REGION Network 241: SAFE OUTPUT CARD FAULT
   RUNG wire#powerrail
      Contact( "reset" )
      { S7_Templates := "SrcType := Word" } EQ_Contact(in1 := "DB101_DB_SDC_FAULTS".Carrier_Fault[7], in2 := 122)
      Coil( "DB302_HMI_Faults".Carrier7_Faults_0.%X9 )
   END_RUNG
   // the same network as SCL:
   "DB302_HMI_Faults".Carrier7_Faults_0.%X9 := "reset" AND ("DB101_DB_SDC_FAULTS".Carrier_Fault[7] = 122);
END_REGION

REGION Network 242: STANDARD INPUT CARD FAULT
   RUNG wire#powerrail
      Contact( "reset" )
      { S7_Templates := "SrcType := Word" } EQ_Contact(in1 := "DB101_DB_SDC_FAULTS".Carrier_Fault[7], in2 := 123)
      Coil( "DB302_HMI_Faults".Carrier7_Faults_0.%X10 )
   END_RUNG
   // the same network as SCL:
   "DB302_HMI_Faults".Carrier7_Faults_0.%X10 := "reset" AND ("DB101_DB_SDC_FAULTS".Carrier_Fault[7] = 123);
END_REGION

REGION Network 243: STANDARD OUTPUT CARD FAULT
   RUNG wire#powerrail
      Contact( "reset" )
      { S7_Templates := "SrcType := Word" } EQ_Contact(in1 := "DB101_DB_SDC_FAULTS".Carrier_Fault[7], in2 := 124)
      Coil( "DB302_HMI_Faults".Carrier7_Faults_0.%X11 )
   END_RUNG
   // the same network as SCL:
   "DB302_HMI_Faults".Carrier7_Faults_0.%X11 := "reset" AND ("DB101_DB_SDC_FAULTS".Carrier_Fault[7] = 124);
END_REGION

REGION Network 244: CARRIER ENCODER POSITION FAULT
   RUNG wire#powerrail
      Contact( "reset" )
      { S7_Templates := "SrcType := Word" } EQ_Contact(in1 := "DB101_DB_SDC_FAULTS".Carrier_Fault[7], in2 := 131)
      Coil( "DB302_HMI_Faults".Carrier7_Faults_0.%X12 )
   END_RUNG
   // the same network as SCL:
   "DB302_HMI_Faults".Carrier7_Faults_0.%X12 := "reset" AND ("DB101_DB_SDC_FAULTS".Carrier_Fault[7] = 131);
END_REGION

REGION Network 245: CARRIER ENCODER INTERNAL ERROR
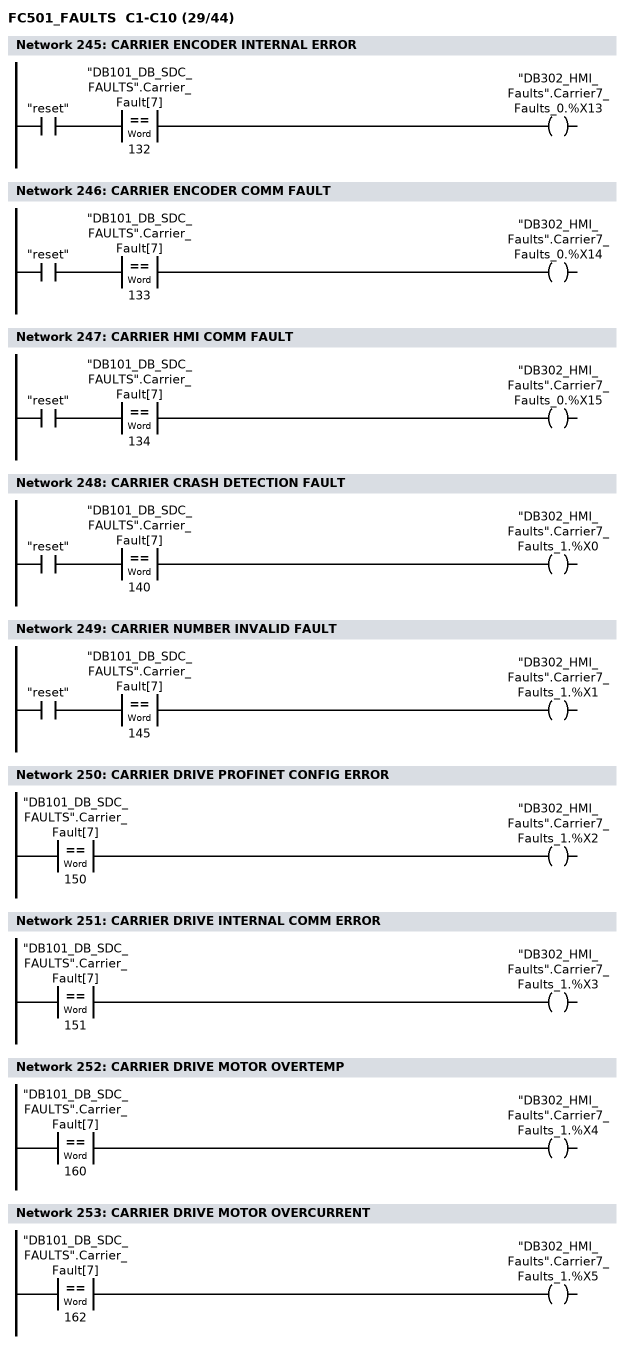
   RUNG wire#powerrail
      Contact( "reset" )
      { S7_Templates := "SrcType := Word" } EQ_Contact(in1 := "DB101_DB_SDC_FAULTS".Carrier_Fault[7], in2 := 132)
      Coil( "DB302_HMI_Faults".Carrier7_Faults_0.%X13 )
   END_RUNG
   // the same network as SCL:
   "DB302_HMI_Faults".Carrier7_Faults_0.%X13 := "reset" AND ("DB101_DB_SDC_FAULTS".Carrier_Fault[7] = 132);
END_REGION

REGION Network 246: CARRIER ENCODER COMM FAULT
   RUNG wire#powerrail
      Contact( "reset" )
      { S7_Templates := "SrcType := Word" } EQ_Contact(in1 := "DB101_DB_SDC_FAULTS".Carrier_Fault[7], in2 := 133)
      Coil( "DB302_HMI_Faults".Carrier7_Faults_0.%X14 )
   END_RUNG
   // the same network as SCL:
   "DB302_HMI_Faults".Carrier7_Faults_0.%X14 := "reset" AND ("DB101_DB_SDC_FAULTS".Carrier_Fault[7] = 133);
END_REGION

REGION Network 247: CARRIER HMI COMM FAULT
   RUNG wire#powerrail
      Contact( "reset" )
      { S7_Templates := "SrcType := Word" } EQ_Contact(in1 := "DB101_DB_SDC_FAULTS".Carrier_Fault[7], in2 := 134)
      Coil( "DB302_HMI_Faults".Carrier7_Faults_0.%X15 )
   END_RUNG
   // the same network as SCL:
   "DB302_HMI_Faults".Carrier7_Faults_0.%X15 := "reset" AND ("DB101_DB_SDC_FAULTS".Carrier_Fault[7] = 134);
END_REGION

REGION Network 248: CARRIER CRASH DETECTION FAULT
   RUNG wire#powerrail
      Contact( "reset" )
      { S7_Templates := "SrcType := Word" } EQ_Contact(in1 := "DB101_DB_SDC_FAULTS".Carrier_Fault[7], in2 := 140)
      Coil( "DB302_HMI_Faults".Carrier7_Faults_1.%X0 )
   END_RUNG
   // the same network as SCL:
   "DB302_HMI_Faults".Carrier7_Faults_1.%X0 := "reset" AND ("DB101_DB_SDC_FAULTS".Carrier_Fault[7] = 140);
END_REGION

REGION Network 249: CARRIER NUMBER INVALID FAULT
   RUNG wire#powerrail
      Contact( "reset" )
      { S7_Templates := "SrcType := Word" } EQ_Contact(in1 := "DB101_DB_SDC_FAULTS".Carrier_Fault[7], in2 := 145)
      Coil( "DB302_HMI_Faults".Carrier7_Faults_1.%X1 )
   END_RUNG
   // the same network as SCL:
   "DB302_HMI_Faults".Carrier7_Faults_1.%X1 := "reset" AND ("DB101_DB_SDC_FAULTS".Carrier_Fault[7] = 145);
END_REGION

REGION Network 250: CARRIER DRIVE PROFINET CONFIG ERROR
   RUNG wire#powerrail
      { S7_Templates := "SrcType := Word" } EQ_Contact(in1 := "DB101_DB_SDC_FAULTS".Carrier_Fault[7], in2 := 150)
      Coil( "DB302_HMI_Faults".Carrier7_Faults_1.%X2 )
   END_RUNG
   // the same network as SCL:
   "DB302_HMI_Faults".Carrier7_Faults_1.%X2 := "DB101_DB_SDC_FAULTS".Carrier_Fault[7] = 150;
END_REGION

REGION Network 251: CARRIER DRIVE INTERNAL COMM ERROR
   RUNG wire#powerrail
      { S7_Templates := "SrcType := Word" } EQ_Contact(in1 := "DB101_DB_SDC_FAULTS".Carrier_Fault[7], in2 := 151)
      Coil( "DB302_HMI_Faults".Carrier7_Faults_1.%X3 )
   END_RUNG
   // the same network as SCL:
   "DB302_HMI_Faults".Carrier7_Faults_1.%X3 := "DB101_DB_SDC_FAULTS".Carrier_Fault[7] = 151;
END_REGION

REGION Network 252: CARRIER DRIVE MOTOR OVERTEMP
   RUNG wire#powerrail
      { S7_Templates := "SrcType := Word" } EQ_Contact(in1 := "DB101_DB_SDC_FAULTS".Carrier_Fault[7], in2 := 160)
      Coil( "DB302_HMI_Faults".Carrier7_Faults_1.%X4 )
   END_RUNG
   // the same network as SCL:
   "DB302_HMI_Faults".Carrier7_Faults_1.%X4 := "DB101_DB_SDC_FAULTS".Carrier_Fault[7] = 160;
END_REGION

REGION Network 253: CARRIER DRIVE MOTOR OVERCURRENT
   RUNG wire#powerrail
      { S7_Templates := "SrcType := Word" } EQ_Contact(in1 := "DB101_DB_SDC_FAULTS".Carrier_Fault[7], in2 := 162)
      Coil( "DB302_HMI_Faults".Carrier7_Faults_1.%X5 )
   END_RUNG
   // the same network as SCL:
   "DB302_HMI_Faults".Carrier7_Faults_1.%X5 := "DB101_DB_SDC_FAULTS".Carrier_Fault[7] = 162;
END_REGION

REGION Network 254: CARRIER DRIVE INFEED OR POWER UNIT NOT READY
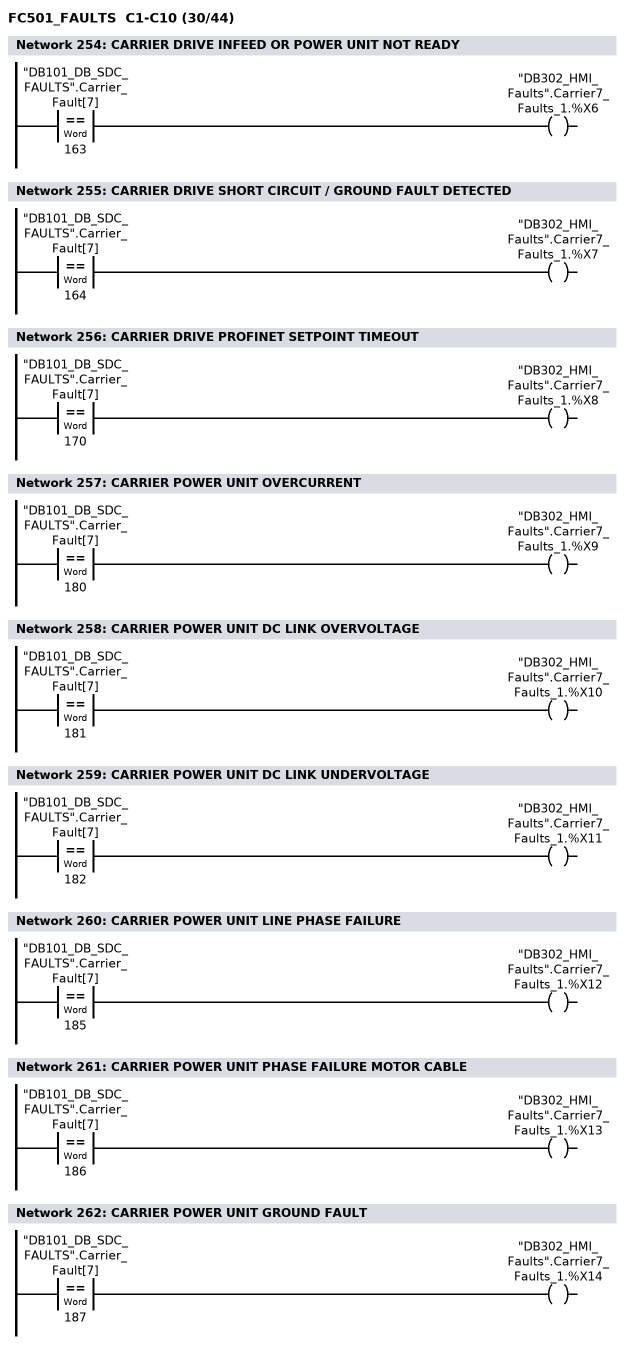
   RUNG wire#powerrail
      { S7_Templates := "SrcType := Word" } EQ_Contact(in1 := "DB101_DB_SDC_FAULTS".Carrier_Fault[7], in2 := 163)
      Coil( "DB302_HMI_Faults".Carrier7_Faults_1.%X6 )
   END_RUNG
   // the same network as SCL:
   "DB302_HMI_Faults".Carrier7_Faults_1.%X6 := "DB101_DB_SDC_FAULTS".Carrier_Fault[7] = 163;
END_REGION

REGION Network 255: CARRIER DRIVE SHORT CIRCUIT / GROUND FAULT DETECTED
   RUNG wire#powerrail
      { S7_Templates := "SrcType := Word" } EQ_Contact(in1 := "DB101_DB_SDC_FAULTS".Carrier_Fault[7], in2 := 164)
      Coil( "DB302_HMI_Faults".Carrier7_Faults_1.%X7 )
   END_RUNG
   // the same network as SCL:
   "DB302_HMI_Faults".Carrier7_Faults_1.%X7 := "DB101_DB_SDC_FAULTS".Carrier_Fault[7] = 164;
END_REGION

REGION Network 256: CARRIER DRIVE PROFINET SETPOINT TIMEOUT
   RUNG wire#powerrail
      { S7_Templates := "SrcType := Word" } EQ_Contact(in1 := "DB101_DB_SDC_FAULTS".Carrier_Fault[7], in2 := 170)
      Coil( "DB302_HMI_Faults".Carrier7_Faults_1.%X8 )
   END_RUNG
   // the same network as SCL:
   "DB302_HMI_Faults".Carrier7_Faults_1.%X8 := "DB101_DB_SDC_FAULTS".Carrier_Fault[7] = 170;
END_REGION

REGION Network 257: CARRIER POWER UNIT OVERCURRENT
   RUNG wire#powerrail
      { S7_Templates := "SrcType := Word" } EQ_Contact(in1 := "DB101_DB_SDC_FAULTS".Carrier_Fault[7], in2 := 180)
      Coil( "DB302_HMI_Faults".Carrier7_Faults_1.%X9 )
   END_RUNG
   // the same network as SCL:
   "DB302_HMI_Faults".Carrier7_Faults_1.%X9 := "DB101_DB_SDC_FAULTS".Carrier_Fault[7] = 180;
END_REGION

REGION Network 258: CARRIER POWER UNIT DC LINK OVERVOLTAGE
   RUNG wire#powerrail
      { S7_Templates := "SrcType := Word" } EQ_Contact(in1 := "DB101_DB_SDC_FAULTS".Carrier_Fault[7], in2 := 181)
      Coil( "DB302_HMI_Faults".Carrier7_Faults_1.%X10 )
   END_RUNG
   // the same network as SCL:
   "DB302_HMI_Faults".Carrier7_Faults_1.%X10 := "DB101_DB_SDC_FAULTS".Carrier_Fault[7] = 181;
END_REGION

REGION Network 259: CARRIER POWER UNIT DC LINK UNDERVOLTAGE
   RUNG wire#powerrail
      { S7_Templates := "SrcType := Word" } EQ_Contact(in1 := "DB101_DB_SDC_FAULTS".Carrier_Fault[7], in2 := 182)
      Coil( "DB302_HMI_Faults".Carrier7_Faults_1.%X11 )
   END_RUNG
   // the same network as SCL:
   "DB302_HMI_Faults".Carrier7_Faults_1.%X11 := "DB101_DB_SDC_FAULTS".Carrier_Fault[7] = 182;
END_REGION

REGION Network 260: CARRIER POWER UNIT LINE PHASE FAILURE
   RUNG wire#powerrail
      { S7_Templates := "SrcType := Word" } EQ_Contact(in1 := "DB101_DB_SDC_FAULTS".Carrier_Fault[7], in2 := 185)
      Coil( "DB302_HMI_Faults".Carrier7_Faults_1.%X12 )
   END_RUNG
   // the same network as SCL:
   "DB302_HMI_Faults".Carrier7_Faults_1.%X12 := "DB101_DB_SDC_FAULTS".Carrier_Fault[7] = 185;
END_REGION

REGION Network 261: CARRIER POWER UNIT PHASE FAILURE MOTOR CABLE
   RUNG wire#powerrail
      { S7_Templates := "SrcType := Word" } EQ_Contact(in1 := "DB101_DB_SDC_FAULTS".Carrier_Fault[7], in2 := 186)
      Coil( "DB302_HMI_Faults".Carrier7_Faults_1.%X13 )
   END_RUNG
   // the same network as SCL:
   "DB302_HMI_Faults".Carrier7_Faults_1.%X13 := "DB101_DB_SDC_FAULTS".Carrier_Fault[7] = 186;
END_REGION

REGION Network 262: CARRIER POWER UNIT GROUND FAULT
   RUNG wire#powerrail
      { S7_Templates := "SrcType := Word" } EQ_Contact(in1 := "DB101_DB_SDC_FAULTS".Carrier_Fault[7], in2 := 187)
      Coil( "DB302_HMI_Faults".Carrier7_Faults_1.%X14 )
   END_RUNG
   // the same network as SCL:
   "DB302_HMI_Faults".Carrier7_Faults_1.%X14 := "DB101_DB_SDC_FAULTS".Carrier_Fault[7] = 187;
END_REGION

REGION Network 263: CARRIER MOTION OFF FAULT
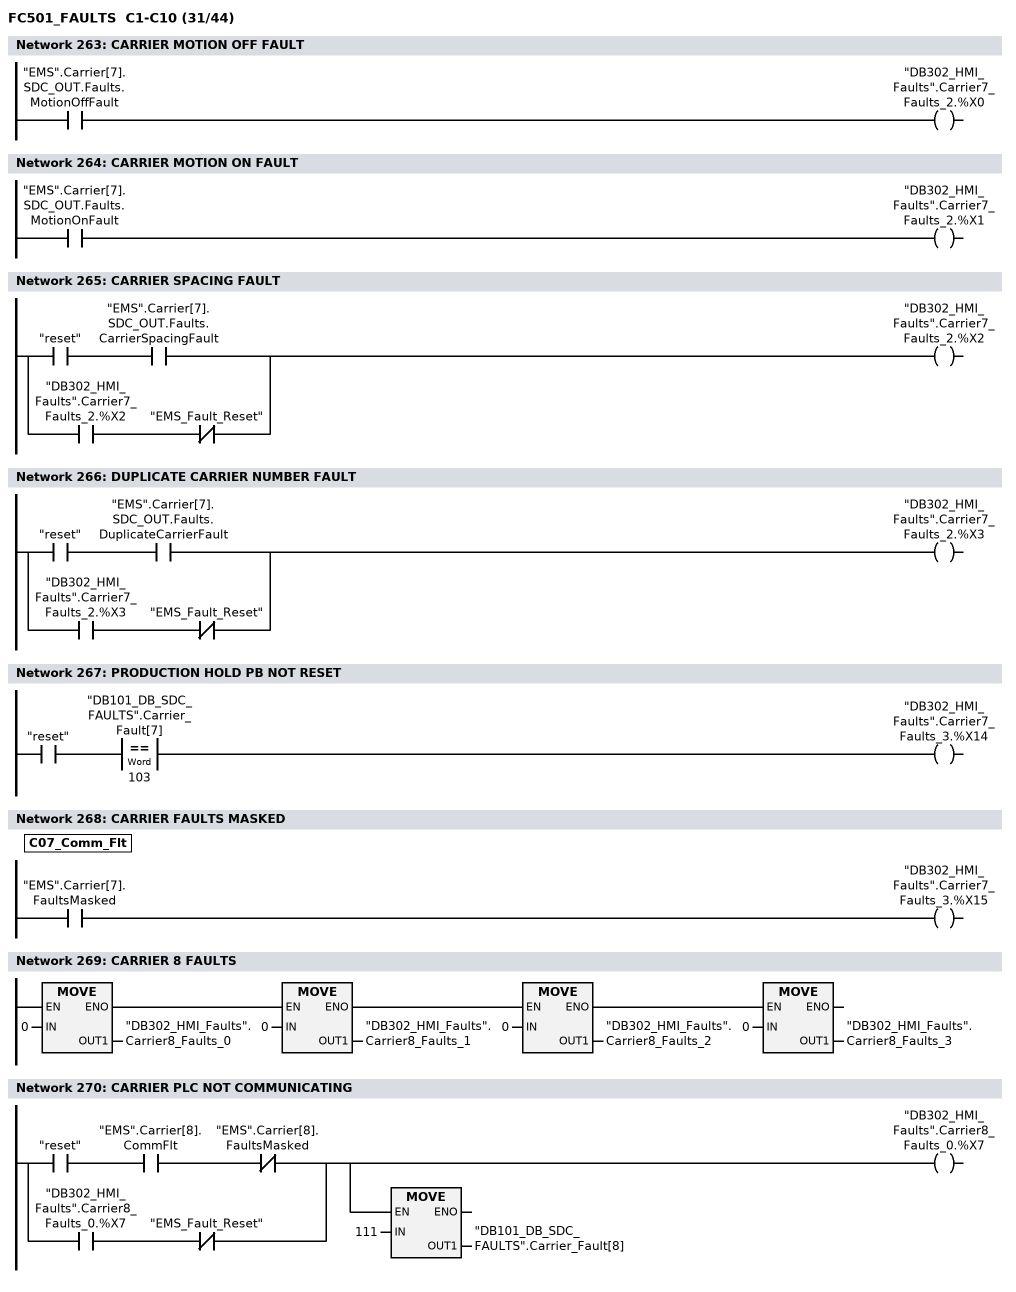
   RUNG wire#powerrail
      Contact( "EMS".Carrier[7].SDC_OUT.Faults.MotionOffFault )
      Coil( "DB302_HMI_Faults".Carrier7_Faults_2.%X0 )
   END_RUNG
   // the same network as SCL:
   "DB302_HMI_Faults".Carrier7_Faults_2.%X0 := "EMS".Carrier[7].SDC_OUT.Faults.MotionOffFault;
END_REGION

REGION Network 264: CARRIER MOTION ON FAULT
   RUNG wire#powerrail
      Contact( "EMS".Carrier[7].SDC_OUT.Faults.MotionOnFault )
      Coil( "DB302_HMI_Faults".Carrier7_Faults_2.%X1 )
   END_RUNG
   // the same network as SCL:
   "DB302_HMI_Faults".Carrier7_Faults_2.%X1 := "EMS".Carrier[7].SDC_OUT.Faults.MotionOnFault;
END_REGION

REGION Network 265: CARRIER SPACING FAULT
   RUNG wire#powerrail
      Contact( "reset" )
      Contact( "EMS".Carrier[7].SDC_OUT.Faults.CarrierSpacingFault )
      wire#w1
      Coil( "DB302_HMI_Faults".Carrier7_Faults_2.%X2 )
   END_RUNG
   RUNG wire#powerrail
      Contact( "DB302_HMI_Faults".Carrier7_Faults_2.%X2 )
      I_Contact( "EMS_Fault_Reset" )
   END_RUNG wire#w1
   // the same network as SCL:
   "DB302_HMI_Faults".Carrier7_Faults_2.%X2 := ("reset" AND "EMS".Carrier[7].SDC_OUT.Faults.CarrierSpacingFault) OR ("DB302_HMI_Faults".Carrier7_Faults_2.%X2 AND NOT "EMS_Fault_Reset");
END_REGION

REGION Network 266: DUPLICATE CARRIER NUMBER FAULT
   RUNG wire#powerrail
      Contact( "reset" )
      Contact( "EMS".Carrier[7].SDC_OUT.Faults.DuplicateCarrierFault )
      wire#w1
      Coil( "DB302_HMI_Faults".Carrier7_Faults_2.%X3 )
   END_RUNG
   RUNG wire#powerrail
      Contact( "DB302_HMI_Faults".Carrier7_Faults_2.%X3 )
      I_Contact( "EMS_Fault_Reset" )
   END_RUNG wire#w1
   // the same network as SCL:
   "DB302_HMI_Faults".Carrier7_Faults_2.%X3 := ("reset" AND "EMS".Carrier[7].SDC_OUT.Faults.DuplicateCarrierFault) OR ("DB302_HMI_Faults".Carrier7_Faults_2.%X3 AND NOT "EMS_Fault_Reset");
END_REGION

REGION Network 267: PRODUCTION HOLD PB NOT RESET
   RUNG wire#powerrail
      Contact( "reset" )
      { S7_Templates := "SrcType := Word" } EQ_Contact(in1 := "DB101_DB_SDC_FAULTS".Carrier_Fault[7], in2 := 103)
      Coil( "DB302_HMI_Faults".Carrier7_Faults_3.%X14 )
   END_RUNG
   // the same network as SCL:
   "DB302_HMI_Faults".Carrier7_Faults_3.%X14 := "reset" AND ("DB101_DB_SDC_FAULTS".Carrier_Fault[7] = 103);
END_REGION

REGION Network 268: CARRIER FAULTS MASKED
   Label( C07_Comm_Flt )
   RUNG wire#powerrail
      Contact( "EMS".Carrier[7].FaultsMasked )
      Coil( "DB302_HMI_Faults".Carrier7_Faults_3.%X15 )
   END_RUNG
   // the same network as SCL:
   C07_Comm_Flt:
   "DB302_HMI_Faults".Carrier7_Faults_3.%X15 := "EMS".Carrier[7].FaultsMasked;
END_REGION

REGION Network 269: CARRIER 8 FAULTS
   RUNG wire#powerrail
      Move(in := 0, out1 => "DB302_HMI_Faults".Carrier8_Faults_0)
      Move(in := 0, out1 => "DB302_HMI_Faults".Carrier8_Faults_1)
      Move(in := 0, out1 => "DB302_HMI_Faults".Carrier8_Faults_2)
      Move(in := 0, out1 => "DB302_HMI_Faults".Carrier8_Faults_3)
   END_RUNG
   // the same network as SCL:
   "DB302_HMI_Faults".Carrier8_Faults_0 := 0;
   "DB302_HMI_Faults".Carrier8_Faults_1 := 0;
   "DB302_HMI_Faults".Carrier8_Faults_2 := 0;
   "DB302_HMI_Faults".Carrier8_Faults_3 := 0;
END_REGION

REGION Network 270: CARRIER PLC NOT COMMUNICATING
   RUNG wire#powerrail
      Contact( "reset" )
      Contact( "EMS".Carrier[8].CommFlt )
      I_Contact( "EMS".Carrier[8].FaultsMasked )
      wire#w1
      Coil( "DB302_HMI_Faults".Carrier8_Faults_0.%X7 )
   END_RUNG
   RUNG wire#powerrail
      Contact( "DB302_HMI_Faults".Carrier8_Faults_0.%X7 )
      I_Contact( "EMS_Fault_Reset" )
   END_RUNG wire#w1
   RUNG wire#w1
      Move(in := 111, out1 => "DB101_DB_SDC_FAULTS".Carrier_Fault[8])
   END_RUNG
   // the same network as SCL:
   "DB302_HMI_Faults".Carrier8_Faults_0.%X7 := ("reset" AND "EMS".Carrier[8].CommFlt AND NOT "EMS".Carrier[8].FaultsMasked) OR ("DB302_HMI_Faults".Carrier8_Faults_0.%X7 AND NOT "EMS_Fault_Reset");
   IF "DB302_HMI_Faults".Carrier8_Faults_0.%X7 THEN "DB101_DB_SDC_FAULTS".Carrier_Fault[8] := 111; END_IF;
END_REGION

REGION Network 271
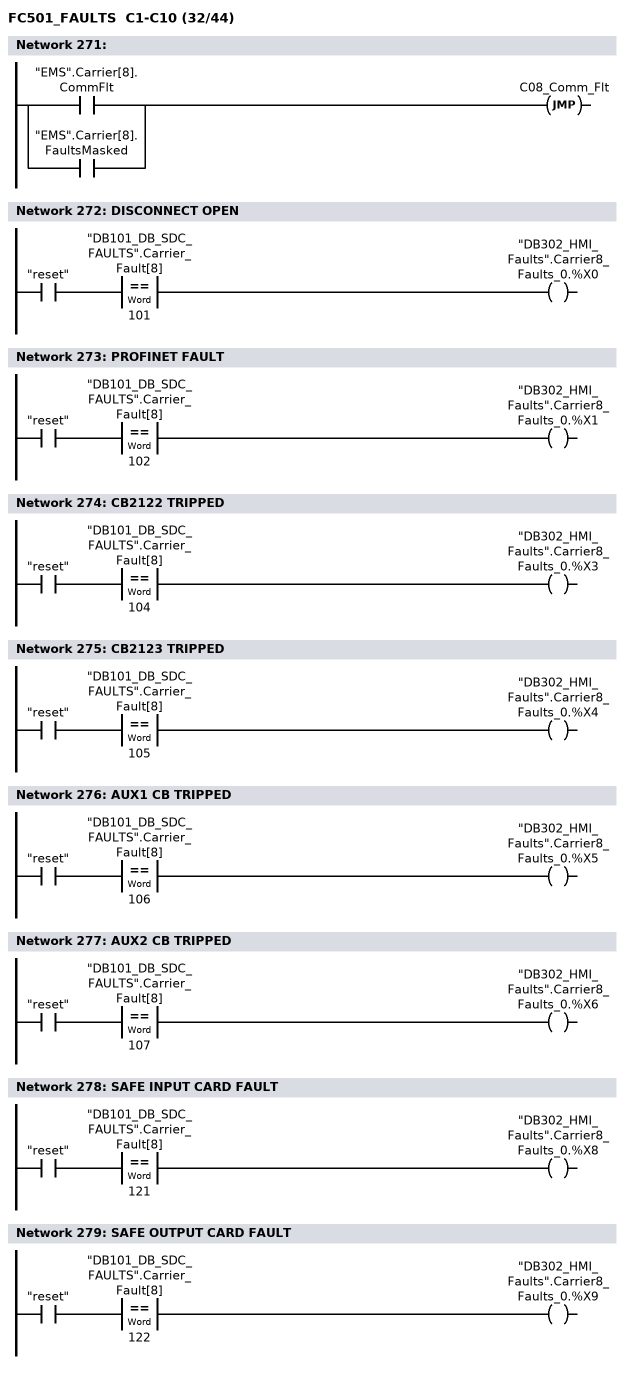
   RUNG wire#powerrail
      Contact( "EMS".Carrier[8].CommFlt )
      wire#w1
      JumpCoil( C08_Comm_Flt )
   END_RUNG
   RUNG wire#powerrail
      Contact( "EMS".Carrier[8].FaultsMasked )
   END_RUNG wire#w1
   // the same network as SCL:
   IF "EMS".Carrier[8].CommFlt OR "EMS".Carrier[8].FaultsMasked THEN GOTO C08_Comm_Flt; END_IF;
END_REGION

REGION Network 272: DISCONNECT OPEN
   RUNG wire#powerrail
      Contact( "reset" )
      { S7_Templates := "SrcType := Word" } EQ_Contact(in1 := "DB101_DB_SDC_FAULTS".Carrier_Fault[8], in2 := 101)
      Coil( "DB302_HMI_Faults".Carrier8_Faults_0.%X0 )
   END_RUNG
   // the same network as SCL:
   "DB302_HMI_Faults".Carrier8_Faults_0.%X0 := "reset" AND ("DB101_DB_SDC_FAULTS".Carrier_Fault[8] = 101);
END_REGION

REGION Network 273: PROFINET FAULT
   RUNG wire#powerrail
      Contact( "reset" )
      { S7_Templates := "SrcType := Word" } EQ_Contact(in1 := "DB101_DB_SDC_FAULTS".Carrier_Fault[8], in2 := 102)
      Coil( "DB302_HMI_Faults".Carrier8_Faults_0.%X1 )
   END_RUNG
   // the same network as SCL:
   "DB302_HMI_Faults".Carrier8_Faults_0.%X1 := "reset" AND ("DB101_DB_SDC_FAULTS".Carrier_Fault[8] = 102);
END_REGION

REGION Network 274: CB2122 TRIPPED
   RUNG wire#powerrail
      Contact( "reset" )
      { S7_Templates := "SrcType := Word" } EQ_Contact(in1 := "DB101_DB_SDC_FAULTS".Carrier_Fault[8], in2 := 104)
      Coil( "DB302_HMI_Faults".Carrier8_Faults_0.%X3 )
   END_RUNG
   // the same network as SCL:
   "DB302_HMI_Faults".Carrier8_Faults_0.%X3 := "reset" AND ("DB101_DB_SDC_FAULTS".Carrier_Fault[8] = 104);
END_REGION

REGION Network 275: CB2123 TRIPPED
   RUNG wire#powerrail
      Contact( "reset" )
      { S7_Templates := "SrcType := Word" } EQ_Contact(in1 := "DB101_DB_SDC_FAULTS".Carrier_Fault[8], in2 := 105)
      Coil( "DB302_HMI_Faults".Carrier8_Faults_0.%X4 )
   END_RUNG
   // the same network as SCL:
   "DB302_HMI_Faults".Carrier8_Faults_0.%X4 := "reset" AND ("DB101_DB_SDC_FAULTS".Carrier_Fault[8] = 105);
END_REGION

REGION Network 276: AUX1 CB TRIPPED
   RUNG wire#powerrail
      Contact( "reset" )
      { S7_Templates := "SrcType := Word" } EQ_Contact(in1 := "DB101_DB_SDC_FAULTS".Carrier_Fault[8], in2 := 106)
      Coil( "DB302_HMI_Faults".Carrier8_Faults_0.%X5 )
   END_RUNG
   // the same network as SCL:
   "DB302_HMI_Faults".Carrier8_Faults_0.%X5 := "reset" AND ("DB101_DB_SDC_FAULTS".Carrier_Fault[8] = 106);
END_REGION

REGION Network 277: AUX2 CB TRIPPED
   RUNG wire#powerrail
      Contact( "reset" )
      { S7_Templates := "SrcType := Word" } EQ_Contact(in1 := "DB101_DB_SDC_FAULTS".Carrier_Fault[8], in2 := 107)
      Coil( "DB302_HMI_Faults".Carrier8_Faults_0.%X6 )
   END_RUNG
   // the same network as SCL:
   "DB302_HMI_Faults".Carrier8_Faults_0.%X6 := "reset" AND ("DB101_DB_SDC_FAULTS".Carrier_Fault[8] = 107);
END_REGION

REGION Network 278: SAFE INPUT CARD FAULT
   RUNG wire#powerrail
      Contact( "reset" )
      { S7_Templates := "SrcType := Word" } EQ_Contact(in1 := "DB101_DB_SDC_FAULTS".Carrier_Fault[8], in2 := 121)
      Coil( "DB302_HMI_Faults".Carrier8_Faults_0.%X8 )
   END_RUNG
   // the same network as SCL:
   "DB302_HMI_Faults".Carrier8_Faults_0.%X8 := "reset" AND ("DB101_DB_SDC_FAULTS".Carrier_Fault[8] = 121);
END_REGION

REGION Network 279: SAFE OUTPUT CARD FAULT
   RUNG wire#powerrail
      Contact( "reset" )
      { S7_Templates := "SrcType := Word" } EQ_Contact(in1 := "DB101_DB_SDC_FAULTS".Carrier_Fault[8], in2 := 122)
      Coil( "DB302_HMI_Faults".Carrier8_Faults_0.%X9 )
   END_RUNG
   // the same network as SCL:
   "DB302_HMI_Faults".Carrier8_Faults_0.%X9 := "reset" AND ("DB101_DB_SDC_FAULTS".Carrier_Fault[8] = 122);
END_REGION

REGION Network 280: STANDARD INPUT CARD FAULT
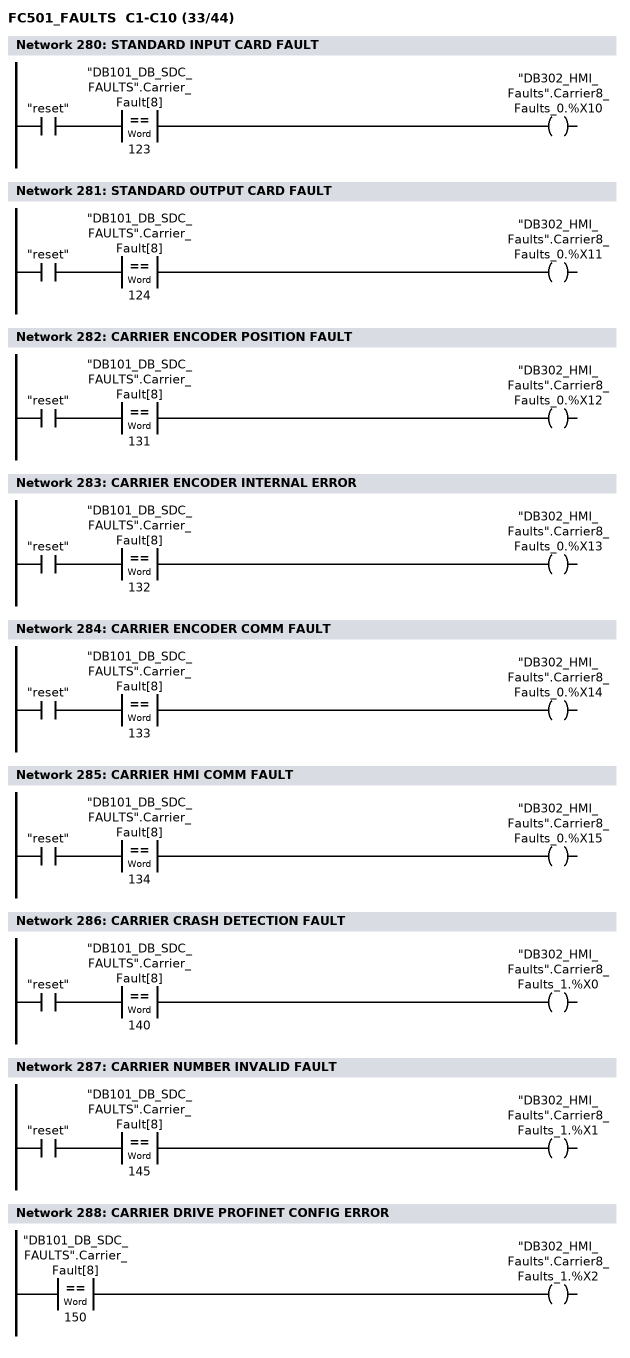
   RUNG wire#powerrail
      Contact( "reset" )
      { S7_Templates := "SrcType := Word" } EQ_Contact(in1 := "DB101_DB_SDC_FAULTS".Carrier_Fault[8], in2 := 123)
      Coil( "DB302_HMI_Faults".Carrier8_Faults_0.%X10 )
   END_RUNG
   // the same network as SCL:
   "DB302_HMI_Faults".Carrier8_Faults_0.%X10 := "reset" AND ("DB101_DB_SDC_FAULTS".Carrier_Fault[8] = 123);
END_REGION

REGION Network 281: STANDARD OUTPUT CARD FAULT
   RUNG wire#powerrail
      Contact( "reset" )
      { S7_Templates := "SrcType := Word" } EQ_Contact(in1 := "DB101_DB_SDC_FAULTS".Carrier_Fault[8], in2 := 124)
      Coil( "DB302_HMI_Faults".Carrier8_Faults_0.%X11 )
   END_RUNG
   // the same network as SCL:
   "DB302_HMI_Faults".Carrier8_Faults_0.%X11 := "reset" AND ("DB101_DB_SDC_FAULTS".Carrier_Fault[8] = 124);
END_REGION

REGION Network 282: CARRIER ENCODER POSITION FAULT
   RUNG wire#powerrail
      Contact( "reset" )
      { S7_Templates := "SrcType := Word" } EQ_Contact(in1 := "DB101_DB_SDC_FAULTS".Carrier_Fault[8], in2 := 131)
      Coil( "DB302_HMI_Faults".Carrier8_Faults_0.%X12 )
   END_RUNG
   // the same network as SCL:
   "DB302_HMI_Faults".Carrier8_Faults_0.%X12 := "reset" AND ("DB101_DB_SDC_FAULTS".Carrier_Fault[8] = 131);
END_REGION

REGION Network 283: CARRIER ENCODER INTERNAL ERROR
   RUNG wire#powerrail
      Contact( "reset" )
      { S7_Templates := "SrcType := Word" } EQ_Contact(in1 := "DB101_DB_SDC_FAULTS".Carrier_Fault[8], in2 := 132)
      Coil( "DB302_HMI_Faults".Carrier8_Faults_0.%X13 )
   END_RUNG
   // the same network as SCL:
   "DB302_HMI_Faults".Carrier8_Faults_0.%X13 := "reset" AND ("DB101_DB_SDC_FAULTS".Carrier_Fault[8] = 132);
END_REGION

REGION Network 284: CARRIER ENCODER COMM FAULT
   RUNG wire#powerrail
      Contact( "reset" )
      { S7_Templates := "SrcType := Word" } EQ_Contact(in1 := "DB101_DB_SDC_FAULTS".Carrier_Fault[8], in2 := 133)
      Coil( "DB302_HMI_Faults".Carrier8_Faults_0.%X14 )
   END_RUNG
   // the same network as SCL:
   "DB302_HMI_Faults".Carrier8_Faults_0.%X14 := "reset" AND ("DB101_DB_SDC_FAULTS".Carrier_Fault[8] = 133);
END_REGION

REGION Network 285: CARRIER HMI COMM FAULT
   RUNG wire#powerrail
      Contact( "reset" )
      { S7_Templates := "SrcType := Word" } EQ_Contact(in1 := "DB101_DB_SDC_FAULTS".Carrier_Fault[8], in2 := 134)
      Coil( "DB302_HMI_Faults".Carrier8_Faults_0.%X15 )
   END_RUNG
   // the same network as SCL:
   "DB302_HMI_Faults".Carrier8_Faults_0.%X15 := "reset" AND ("DB101_DB_SDC_FAULTS".Carrier_Fault[8] = 134);
END_REGION

REGION Network 286: CARRIER CRASH DETECTION FAULT
   RUNG wire#powerrail
      Contact( "reset" )
      { S7_Templates := "SrcType := Word" } EQ_Contact(in1 := "DB101_DB_SDC_FAULTS".Carrier_Fault[8], in2 := 140)
      Coil( "DB302_HMI_Faults".Carrier8_Faults_1.%X0 )
   END_RUNG
   // the same network as SCL:
   "DB302_HMI_Faults".Carrier8_Faults_1.%X0 := "reset" AND ("DB101_DB_SDC_FAULTS".Carrier_Fault[8] = 140);
END_REGION

REGION Network 287: CARRIER NUMBER INVALID FAULT
   RUNG wire#powerrail
      Contact( "reset" )
      { S7_Templates := "SrcType := Word" } EQ_Contact(in1 := "DB101_DB_SDC_FAULTS".Carrier_Fault[8], in2 := 145)
      Coil( "DB302_HMI_Faults".Carrier8_Faults_1.%X1 )
   END_RUNG
   // the same network as SCL:
   "DB302_HMI_Faults".Carrier8_Faults_1.%X1 := "reset" AND ("DB101_DB_SDC_FAULTS".Carrier_Fault[8] = 145);
END_REGION

REGION Network 288: CARRIER DRIVE PROFINET CONFIG ERROR
   RUNG wire#powerrail
      { S7_Templates := "SrcType := Word" } EQ_Contact(in1 := "DB101_DB_SDC_FAULTS".Carrier_Fault[8], in2 := 150)
      Coil( "DB302_HMI_Faults".Carrier8_Faults_1.%X2 )
   END_RUNG
   // the same network as SCL:
   "DB302_HMI_Faults".Carrier8_Faults_1.%X2 := "DB101_DB_SDC_FAULTS".Carrier_Fault[8] = 150;
END_REGION

REGION Network 289: CARRIER DRIVE INTERNAL COMM ERROR
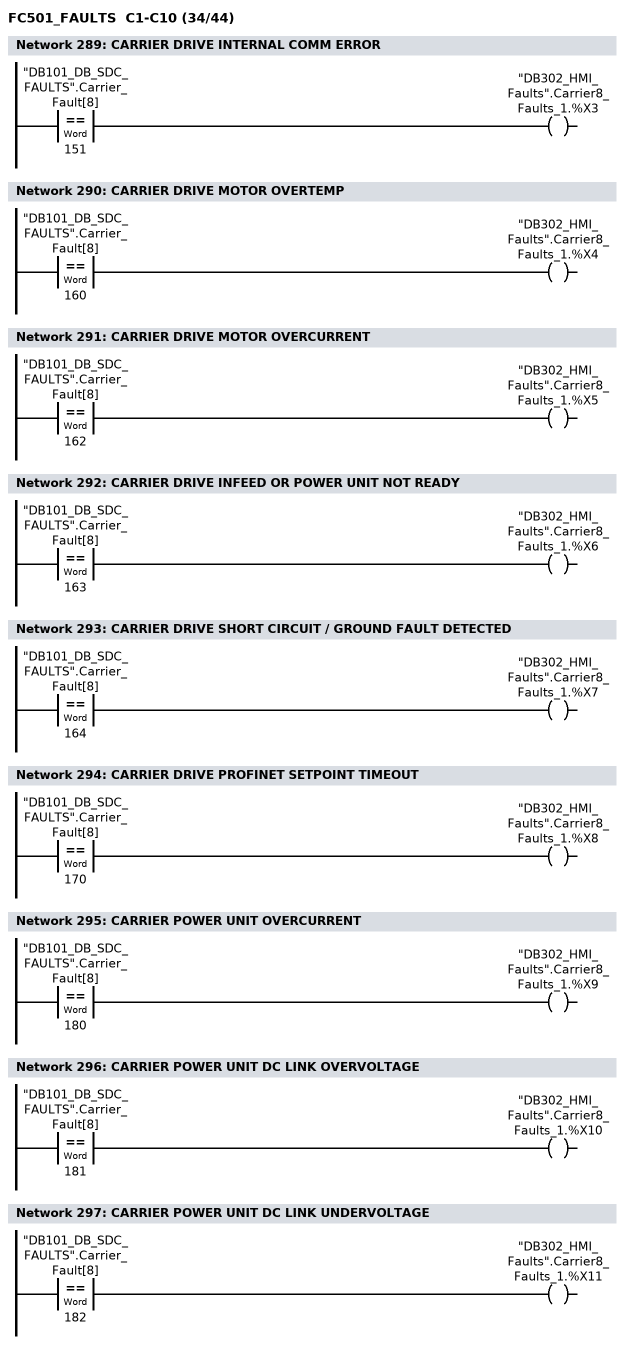
   RUNG wire#powerrail
      { S7_Templates := "SrcType := Word" } EQ_Contact(in1 := "DB101_DB_SDC_FAULTS".Carrier_Fault[8], in2 := 151)
      Coil( "DB302_HMI_Faults".Carrier8_Faults_1.%X3 )
   END_RUNG
   // the same network as SCL:
   "DB302_HMI_Faults".Carrier8_Faults_1.%X3 := "DB101_DB_SDC_FAULTS".Carrier_Fault[8] = 151;
END_REGION

REGION Network 290: CARRIER DRIVE MOTOR OVERTEMP
   RUNG wire#powerrail
      { S7_Templates := "SrcType := Word" } EQ_Contact(in1 := "DB101_DB_SDC_FAULTS".Carrier_Fault[8], in2 := 160)
      Coil( "DB302_HMI_Faults".Carrier8_Faults_1.%X4 )
   END_RUNG
   // the same network as SCL:
   "DB302_HMI_Faults".Carrier8_Faults_1.%X4 := "DB101_DB_SDC_FAULTS".Carrier_Fault[8] = 160;
END_REGION

REGION Network 291: CARRIER DRIVE MOTOR OVERCURRENT
   RUNG wire#powerrail
      { S7_Templates := "SrcType := Word" } EQ_Contact(in1 := "DB101_DB_SDC_FAULTS".Carrier_Fault[8], in2 := 162)
      Coil( "DB302_HMI_Faults".Carrier8_Faults_1.%X5 )
   END_RUNG
   // the same network as SCL:
   "DB302_HMI_Faults".Carrier8_Faults_1.%X5 := "DB101_DB_SDC_FAULTS".Carrier_Fault[8] = 162;
END_REGION

REGION Network 292: CARRIER DRIVE INFEED OR POWER UNIT NOT READY
   RUNG wire#powerrail
      { S7_Templates := "SrcType := Word" } EQ_Contact(in1 := "DB101_DB_SDC_FAULTS".Carrier_Fault[8], in2 := 163)
      Coil( "DB302_HMI_Faults".Carrier8_Faults_1.%X6 )
   END_RUNG
   // the same network as SCL:
   "DB302_HMI_Faults".Carrier8_Faults_1.%X6 := "DB101_DB_SDC_FAULTS".Carrier_Fault[8] = 163;
END_REGION

REGION Network 293: CARRIER DRIVE SHORT CIRCUIT / GROUND FAULT DETECTED
   RUNG wire#powerrail
      { S7_Templates := "SrcType := Word" } EQ_Contact(in1 := "DB101_DB_SDC_FAULTS".Carrier_Fault[8], in2 := 164)
      Coil( "DB302_HMI_Faults".Carrier8_Faults_1.%X7 )
   END_RUNG
   // the same network as SCL:
   "DB302_HMI_Faults".Carrier8_Faults_1.%X7 := "DB101_DB_SDC_FAULTS".Carrier_Fault[8] = 164;
END_REGION

REGION Network 294: CARRIER DRIVE PROFINET SETPOINT TIMEOUT
   RUNG wire#powerrail
      { S7_Templates := "SrcType := Word" } EQ_Contact(in1 := "DB101_DB_SDC_FAULTS".Carrier_Fault[8], in2 := 170)
      Coil( "DB302_HMI_Faults".Carrier8_Faults_1.%X8 )
   END_RUNG
   // the same network as SCL:
   "DB302_HMI_Faults".Carrier8_Faults_1.%X8 := "DB101_DB_SDC_FAULTS".Carrier_Fault[8] = 170;
END_REGION

REGION Network 295: CARRIER POWER UNIT OVERCURRENT
   RUNG wire#powerrail
      { S7_Templates := "SrcType := Word" } EQ_Contact(in1 := "DB101_DB_SDC_FAULTS".Carrier_Fault[8], in2 := 180)
      Coil( "DB302_HMI_Faults".Carrier8_Faults_1.%X9 )
   END_RUNG
   // the same network as SCL:
   "DB302_HMI_Faults".Carrier8_Faults_1.%X9 := "DB101_DB_SDC_FAULTS".Carrier_Fault[8] = 180;
END_REGION

REGION Network 296: CARRIER POWER UNIT DC LINK OVERVOLTAGE
   RUNG wire#powerrail
      { S7_Templates := "SrcType := Word" } EQ_Contact(in1 := "DB101_DB_SDC_FAULTS".Carrier_Fault[8], in2 := 181)
      Coil( "DB302_HMI_Faults".Carrier8_Faults_1.%X10 )
   END_RUNG
   // the same network as SCL:
   "DB302_HMI_Faults".Carrier8_Faults_1.%X10 := "DB101_DB_SDC_FAULTS".Carrier_Fault[8] = 181;
END_REGION
